   "DB_Integer_IHour" : USInt = PLC Data_Integer.IHour, 1 s
   "DB_Integer_IMinute" : USInt = PLC Data_Integer.IMinute, 1 s
   "DB_Integer_IMonth" : USInt = PLC Data_Integer.IMonth, 1 s
   "DB_Integer_ISecond" : USInt = PLC Data_Integer.ISecond, 1 s
   "DB_Integer_IYear" : UInt = PLC Data_Integer.IYear, 1 s
   "DB_Integer_S1AHour" : USInt = PLC Data_Integer.S1AHour, 1 s
   "DB_Integer_S1AMinute" : USInt = PLC Data_Integer.S1AMinute, 1 s
   "DB_Integer_S1ASecond" : USInt = PLC Data_Integer.S1ASecond, 1 s
   "DB_Integer_S1BHour" : USInt = PLC Data_Integer.S1BHour, 1 s
   "DB_Integer_S1BMinute" : USInt = PLC Data_Integer.S1BMinute, 1 s
   "DB_Integer_S1BSecond" : USInt = PLC Data_Integer.S1BSecond, 1 s
   "DB_Integer_S2AHour" : USInt = PLC Data_Integer.S2AHour, 1 s
   "DB_Integer_S2AMinute" : USInt = PLC Data_Integer.S2AMinute, 1 s
   "DB_Integer_S2ASecond" : USInt = PLC Data_Integer.S2ASecond, 1 s
   "DB_Integer_S2BHour" : USInt = PLC Data_Integer.S2BHour, 1 s
   "DB_Integer_S2BMinute" : USInt = PLC Data_Integer.S2BMinute, 1 s
   "DB_Integer_S2BSecond" : USInt = PLC Data_Integer.S2BSecond, 1 s
   "DB_Integer_S3AHour" : USInt = PLC Data_Integer.S3AHour, 1 s
   "DB_Integer_S3AMinute" : USInt = PLC Data_Integer.S3AMinute, 1 s
   "DB_Integer_S3ASecond" : USInt = PLC Data_Integer.S3ASecond, 1 s
   "DB_Integer_S3BHour" : USInt = PLC Data_Integer.S3BHour, 1 s
   "DB_Integer_S3BMinute" : USInt = PLC Data_Integer.S3BMinute, 1 s
   "DB_Integer_S3BSecond" : USInt = PLC Data_Integer.S3BSecond, 1 s
   "DB_Real_% Reject Out Stop[0]" : Real = PLC Data_Real."% Reject Out Stop"[0], 1 s
   "DB_Real_% Reject Out Stop[1]" : Real = PLC Data_Real."% Reject Out Stop"[1], 1 s
   "DB_Real_% Reject Out Stop[2]" : Real = PLC Data_Real."% Reject Out Stop"[2], 1 s
   "DB_Real_% Reject Out Stop[3]" : Real = PLC Data_Real."% Reject Out Stop"[3], 1 s
   "DB_Real_% Reject Out Stop[4]" : Real = PLC Data_Real."% Reject Out Stop"[4], 1 s
   "DB_Real_% Reject Out Stop[5]" : Real = PLC Data_Real."% Reject Out Stop"[5], 1 s
   "DB_Real_%Bad Read" : Array [0..5] of Real = PLC Data_Real."%Bad Read", 1 s
   "DB_Real_%Bad Read[0]" : Real = PLC Data_Real."%Bad Read"[0], 1 s
   "DB_Real_%Bad Read[1]" : Real = PLC Data_Real."%Bad Read"[1], 1 s
   "DB_Real_%Bad Read[2]" : Real = PLC Data_Real."%Bad Read"[2], 1 s
   "DB_Real_%Bad Read[3]" : Real = PLC Data_Real."%Bad Read"[3], 1 s
   "DB_Real_%Bad Read[4]" : Real = PLC Data_Real."%Bad Read"[4], 1 s
   "DB_Real_%Bad Read[5]" : Real = PLC Data_Real."%Bad Read"[5], 1 s
   "DB_Real_%Good Read[0]" : Real = PLC Data_Real."%Good Read"[0], 1 s
   "DB_Real_%Good Read[1]" : Real = PLC Data_Real."%Good Read"[1], 1 s
   "DB_Real_%Good Read[2]" : Real = PLC Data_Real."%Good Read"[2], 1 s
   "DB_Real_%Good Read[3]" : Real = PLC Data_Real."%Good Read"[3], 1 s
   "DB_Real_%Good Read[4]" : Real = PLC Data_Real."%Good Read"[4], 1 s
   "DB_Real_%Good Read[5]" : Real = PLC Data_Real."%Good Read"[5], 1 s
   "DB_Real_Efficiency CS" : Array [0..5] of Real = PLC Data_Real."% Reject Out Stop", 1 s

discrete alarms
   1: 'Pressure Low', class Errors, trigger "HMI_Tag_1" bit 8
   2: 'Door Open Labelling', class Errors, trigger "HMI_Tag_1" bit 9
   3: 'Door Open Focke Chute', class Errors, trigger "HMI_Tag_1" bit 10
   4: 'Chute 3 Way Full', class Errors, trigger "HMI_Tag_1" bit 11
   5: 'Door Open FC Proximity', class Errors, trigger "HMI_Tag_1" bit 12
   6: 'Alarm2', class Errors, trigger "HMI_Tag_1" bit 13
   7: 'Imaje Paper/Ribbon Out', class Errors, trigger "HMI_Tag_1" bit 14
   8: 'Imaje System Error', class Errors, trigger "HMI_Tag_1" bit 15
   9: 'Imaje Not In Position', class Errors, trigger "HMI_Tag_1" bit 0
   10: 'Heater Not Ready', class Errors, trigger "HMI_Tag_1" bit 1
   11: 'Reed Switch Pneumatic 1 Pusher', class Errors, trigger "HMI_Tag_1" bit 2
   12: 'Alarm3', class Errors, trigger "HMI_Tag_1" bit 3
   13: 'Reed Switch Pneumatic 3 Up', class Errors, trigger "HMI_Tag_1" bit 4
   14: 'Reed Switch Pneumatic 3 Down', class Errors, trigger "HMI_Tag_1" bit 5
   15: 'Reed Switch Pneumatic 4 Down', class Errors, trigger "HMI_Error_Cont" bit 8
   16: 'Reed Switch Pneumatic 4 Up', class Errors, trigger "HMI_Error_Cont" bit 9
   17: 'Reed Switch Pneumatic 5 Advance', class Errors, trigger "HMI_Error_Cont" bit 10
   18: 'Reed Switch Pneumatic 5 Retract', class Errors, trigger "HMI_Error_Cont" bit 11
   19: 'Chute Heating Roll Full', class Errors, trigger "HMI_Tag_1" bit 6

text list "Machine Running": 0 'STOP'; 1 'RUNNING'

text list "Status Markem": 0 'PAUSE'; 1 'START'

text list "Mode Machine": 0 'With Focke Chute'; 1 'Without Focke Chute'

text list "Mode Bypass": 0 'OFF'; 1 'ON'

Template "Template_1" 320x240
   Button "Template_" at 267,190 size 51x47; TextOff 'ExitRuntime'; PictureOff "ExitRuntime_HMI_1"; PictureOn "ExitRuntime_HMI_1"
      on Release: StopRuntime(0)
   Button "Template_1" at 214,190 size 51x47; TextOff 'Text'
   Button "Template_2" at 160,190 size 51x47; TextOff 'Text'
   Button "Template_3" at 107,190 size 51x47; TextOff 'Login'; PictureOff "Login_HMI_1"; PictureOn "Login_HMI_1"
      on Release: function_a2a04561()
   Button "Template_4" at 54,190 size 51x47; TextOff 'AlarmDisplay'; PictureOff "AlarmDisplay_HMI_1"; PictureOn "AlarmDisplay_HMI_1"
      on Release: function_ef3f5d25("Alarm window_Unacknowledged", -1)
   Button "Template_5" at 1,190 size 51x47; TextOff 'NavigateHome'; PictureOff "NavigateHome_HMI_1"; PictureOn "NavigateHome_HMI_1"
   SymbolicIOField "Symbolic_IO_Field_Screen" at 73,7 size 160x25; TextOff '0'; TextOn '1'; TextList "TextList_ScreenNames"
      ProcessValue <- "Tag_ScreenNumber"
   DateTimeField "Template_6" at 235,20 size 85x20
   DateTimeField "Template_7" at 235,0 size 85x20
   GraphicView "Logo" at 0,0 size 71x40; Picture "Logo of HMI_1"

screen "Introduction" 320x240
   Button "Button_1" at 100,200 size 120x30; TextOff 'Go to Main Page'
      on Click: ActivateScreen("Main Page", 0)
   GraphicView "Graphic view_1" at 0,0 size 319x37; Picture "Logo SMS"
   TextField "Text field_1" at 6,54 size 278x31; Text 'END LABELLER MACHINE'
   TextField "Text field_2" at 19,85 size 278x92; Text 'Production : 65 Slof/minute Electric Power : 2,5 KW Compressed Air : 6 Bar Program Version : 14.6 Year : 2013'

screen "Main Page" 320x240
   on GenerateScreen: SetBit("Flag Main Page")
   TextField "Text field_1" at 106,1 size 113x25; Text 'MAIN PAGE'
   TextField "Text field_3" at 5,50 size 91x15; Text 'Machine Status'
   TextField "Text field_4" at 5,73 size 91x15; Text 'Markem Status'
   SymbolicIOField "Symbolic I/O field_2" at 100,48 size 122x19; TextOff '0'; TextOn '1'; TextList "Machine Running"
      ProcessValue <- "Machine Running"
   SymbolicIOField "Symbolic I/O field_1" at 100,71 size 122x19; TextOff '0'; TextOn '1'; TextList "Status Markem"
      ProcessValue <- "Flag Imaje Start"
   Button "Button_4" at 0,209 size 90x30; TextOff 'Test Mode'
      on Click: ActivateScreen("Test Mode", 0)
   Button "Button_5" at 95,209 size 90x30; TextOff 'Parameter'
      on Click: ActivateScreen("Parameter", 0)
   TextField "Text field_5" at 5,95 size 91x15; Text 'Mode Machine'
   SymbolicIOField "Symbolic I/O field_3" at 100,94 size 122x19; TextOff '0'; TextOn '1'; TextList "Mode Machine"
      ProcessValue <- "Flag Enable/Disable Block Focke"
   TextField "Text field_7" at 5,117 size 91x15; Text 'Mode Bypass'
   SymbolicIOField "Symbolic I/O field_4" at 100,117 size 122x19; TextOff '0'; TextOn '1'; TextList "Mode Bypass"
      ProcessValue <- "Flag Machine Bypass"
   IOField "I/O field_3" at 85,24 size 155x23; FormatPattern 9999999999999999999999999999999999999999
      ProcessValue <- "DB_DTL1_Output"
   Button "Button_1" at 287,1 size 29x23; TextOff 'Text'
      on Click: StopRuntime(0)
   Button "Button_2" at 193,208 size 120x30; TextOff 'Statistika Data'
      on Click: ActivateScreen("Data Statistika", 0)

screen "Parameter" 320x240
   on GenerateScreen: SetBit("Flag Parameter Page")
   on ClearScreen: ResetBit("Flag Parameter Page")
   TextField "Text field_1" at 1,0 size 319x27; Text 'PARAMETER'
   Button "Button_4" at 91,202 size 132x30; TextOff 'Back to Main Page'
      on Click: ActivateScreen("Main Page", 0)
   Button "Button_3" at 91,48 size 132x30; TextOff 'Setting Timer'
      on Click: ActivateScreen("Setting Timer", 0)
   Button "Button_2" at 91,88 size 132x30; TextOff 'Setting Machine'
      on Click: ActivateScreen("Setting Machine", 0)

screen "Setting Timer" 320x240
   on ClearScreen: ResetBit("Flag Parameter Page")
   on GenerateScreen: SetBit("Flag Parameter Page")
   TextField "Text field_1" at 0,0 size 319x27; Text 'SETTING TIMER'
   Button "Button_2" at 92,200 size 120x30; TextOff 'Back to Parameter'
      on Click: ActivateScreen("Parameter", 0)
   TextField "Text field_2" at 5,39 size 150x15; Text 'Timer Delay Stamp'
   IOField "I/O field_1" at 152,40 size 80x16; FormatPattern 9999; Unit  ms
      ProcessValue <- "Timer Delay Stamp"
   TextField "Text field_3" at 5,63 size 150x15; Text 'Timer Scanning Barcode'
   IOField "I/O field_2" at 153,64 size 80x16; FormatPattern 9999; Unit  ms
      ProcessValue <- "Timer Trigger Barcode"

screen "Test Mode" 320x240
   on GenerateScreen: SetBit("PB Test Mode")
   on ClearScreen: ResetBit("PB Test Mode")
   TextField "Text field_1" at 1,1 size 319x27; Text 'TEST MODE'
   Switch "Switch_1" at 3,34 size 95x30; TextOff 'Pneumatic 1 Off'; CaptionText 'Switch'; TextOn 'Pneumatic 1 On'
      ProcessValue <- "PB Test Pneumatic 1"
   Switch "Switch_2" at 3,75 size 95x30; CaptionText 'Switch'; TextOff 'Pneumatic 2 Off'; TextOn 'Pneumatic 2 On'
      ProcessValue <- "PB Test Pneumatic 2"
   Switch "Switch_3" at 3,116 size 95x30; CaptionText 'Switch'; TextOff 'Pneumatic 3 Off'; TextOn 'Pneumatic 3 On'
      ProcessValue <- "PB Test Pneumatic 3"
   Switch "Switch_5" at 104,34 size 115x30; CaptionText 'Switch'; TextOff 'Pneumatic 5 Off'; TextOn 'Pneumatic 5 On'
      ProcessValue <- "PB Test Pneumatic 5"
   Switch "Switch_6" at 226,116 size 90x30; CaptionText 'Switch'; TextOff 'Motor Off'; TextOn 'Motor On'
      ProcessValue <- "PB Test Motor"
   Button "Button_1" at 100,204 size 120x30; TextOff 'Back to Main Page'
      on Click: ActivateScreen("Main Page", 0)
   Button "Button_2" at 226,34 size 90x30; TextOff 'Stamp Off'; TextOn 'Stamp On'
      on Press: SetBit("PB Test Imaje")
      on Release: ResetBit("PB Test Imaje")
   Switch "Switch_7" at 104,116 size 115x30; CaptionText 'Switch'; TextOff 'Air Valve On'; TextOn 'Air Valve Off'
      ProcessValue <- "PB Test Air Valve"
   Button "Button_3" at 226,75 size 90x30; TextOff 'Teach In'
      on Press: SetBit("Flag Teach In Barcode")
      on Release: ResetBit("Flag Teach In Barcode")
   Switch "Switch_8" at 3,157 size 95x30; CaptionText 'Switch'; TextOff 'Pneumatic 4 Off'; TextOn 'Pneumatic 4 On'
      ProcessValue <- "PB Test Pneumatic 4"
   Switch "Switch_4" at 104,75 size 115x30; CaptionText 'Switch'; TextOff 'Pneumatic 6 On'; TextOn 'Pneumatic 6 Off'
      ProcessValue <- "PB Test Pneumatic 6"
   Switch "Switch_9" at 104,157 size 115x30; CaptionText 'Switch'; TextOff 'Conveyor Pusher Off'; TextOn 'Conveyor Pusher On'
      ProcessValue <- "PB Test Motor Coveyor Pusher"
   Switch "Switch_10" at 226,157 size 90x30; CaptionText 'Switch'; TextOff 'Heating Roll Off'; TextOn 'Heating Roll On'
      ProcessValue <- "PB Test Motor Heating Roll"

screen "Setting Machine" 320x240
   on ClearScreen: ResetBit("Flag Parameter Page")
   on GenerateScreen: SetBit("Flag Parameter Page")
   TextField "Text field_1" at 1,0 size 319x27; Text 'SETTING MACHINE'
   Switch "Switch_1" at 16,38 size 135x30; CaptionText 'Switch'; TextOff 'Barcode Off'; TextOn 'Barcode ON'
      ProcessValue <- "Flag Barcode HMI"
   Switch "Switch_2" at 16,108 size 135x30; CaptionText 'Switch'; TextOff 'Chute 3Way Error ON'; TextOn 'Chute 3Way Error OFF'
      ProcessValue <- "Flag Enable/Disable Error Chute 3 Way"
   Button "Button_2" at 101,205 size 120x30; TextOff 'Back to Parameter'
      on Click: ActivateScreen("Parameter", 0)
   Switch "Switch_3" at 16,73 size 135x30; CaptionText 'Switch'; TextOff 'Heater Error Off'; TextOn 'Heater Error ON'
      ProcessValue <- "Flag Heater Error HMI"
   Switch "Switch_4" at 170,38 size 135x30; CaptionText 'Switch'; TextOff 'Reed Switch Bypass Off'; TextOn 'Reed Switch Bypass On'
      ProcessValue <- "Flag Pneumatic Bypass"
   Switch "Switch_5" at 170,108 size 135x30; CaptionText 'Switch'; TextOff 'Safety Door On'; TextOn 'Safety Door Off'
      ProcessValue <- "Flag Enable/Disable Error Door Open"
   Button "Button_1" at 289,0 size 31x30; TextOff 'Setting Mode'; Authorization "User administration"
      on Click: ActivateScreen("Setting Mode", 0)
   Button "Button_3" at 170,73 size 135x30; TextOff 'Setting Reed Switch'
      on Click: ActivateScreen("Setting Reed Switch", 0)
   Switch "Switch_6" at 16,143 size 135x30; CaptionText 'Switch'; TextOff 'Chute Heating Roll Error ON'; TextOn 'Chute Heating Roll Error OFF'
      ProcessValue <- "Flag Enable/Disable Error Chute Before Heating Roll"
   Softkey "Softkey_F6" at 266,202 size 53x38
      on KeyDown: ActivateScreen("Setting Mode", 0)
      on KeyUp: ActivateScreen("Setting Mode", 0)
   Softkey "Softkey_F5" at 213,202 size 53x38
      on KeyDown: function_f23ef4c9()
      on KeyUp: function_f23ef4c9()

screen "Setting Mode" 320x240
   TextField "Text field_1" at 1,0 size 319x27; Text 'MODE MACHINE'
   Button "Button_1" at 95,203 size 129x30; TextOff 'Back to Setting Machine'
      on Click: ActivateScreen("Setting Machine", 0)
   Switch "Switch_1" at 70,46 size 177x32; CaptionText 'Switch'; TextOff 'With Focke Chute'; TextOn 'Without Focke Chute'
      ProcessValue <- "Flag Enable/Disable Block Focke"
   Switch "Switch_2" at 70,90 size 177x32; TextOff 'Disable Flow to Reject'; CaptionText 'Switch'; TextOn 'Enable Flow to Reject'
      ProcessValue <- "Flag Enable/Disable Flow to Reject"
   Switch "Switch_3" at 70,130 size 177x32; TextOff 'With Heating Roll'; CaptionText 'Switch'; TextOn 'Without Heating Roll'
      ProcessValue <- "Flag Enable/Disable Heating Roll"

screen "Setting Reed Switch" 320x240
   TextField "Text field_1" at 1,3 size 319x27; Text 'SETTING REED SWITCH BYPASS'
   Switch "Switch_4" at 21,103 size 128x30; CaptionText 'Switch'; TextOff 'RS Pneu 3 Bypass Off'; TextOn 'RS Pneu 3 Bypass On'
      ProcessValue <- "RS Bypass Pneumatic 3"
   Switch "Switch_1" at 172,103 size 128x30; CaptionText 'Switch'; TextOff 'RS Pneu 5 Bypass Off'; TextOn 'RS Pneu 5 Bypass On'
      ProcessValue <- "RS Bypass Pneumatic 5"
   Switch "Switch_2" at 172,59 size 128x30; CaptionText 'Switch'; TextOff 'RS Pneu 4 Bypass Off'; TextOn 'RS Pneu 4 Bypass On'
      ProcessValue <- "RS Bypass Pneumatic 4"
   Switch "Switch_3" at 21,59 size 128x30; CaptionText 'Switch'; TextOff 'RS Pneu 1 Bypass Off'; TextOn 'RS Pneu 1 Bypass On'
      ProcessValue <- "RS Bypass Pneumatic 1"
   Button "Button_1" at 95,203 size 129x30; TextOff 'Back to Setting Machine'
      on Click: ActivateScreen("Setting Machine", 0)

screen "Data Current Shift" 320x240
   IOField "I/O field_11" at 221,82 size 60x19; FormatPattern 999.99; Unit   %
      ProcessValue <- "Data_Real_% Total Output[0]"
   IOField "I/O field_9" at 221,102 size 60x19; FormatPattern 999.99; Unit   %
      ProcessValue <- "DB_Real_%Good Read[0]"
   IOField "I/O field_8" at 221,120 size 60x19; FormatPattern 999.99; Unit   %
      ProcessValue <- "DB_Real_%Bad Read[0]"
   TextField "Text field_1" at 92,0 size 137x18; Text 'CURRENT SHIFT DATA'
   IOField "I/O field_1" at 142,59 size 79x19; FormatPattern 99999999; Unit  Pcs
      ProcessValue <- "DB_IntData_Input Sloft"
   TextField "Text field_2" at 4,60 size 138x17; Text 'Input Sloft'
   TextField "Text field_3" at 4,83 size 138x17; Text 'Total Output Sloft'
   TextField "Text field_4" at 4,101 size 138x19; Text 'Good Read Sloft'
   TextField "Text field_7" at 4,121 size 138x18; Text 'Bad Read Sloft'
   IOField "I/O field_3" at 142,101 size 79x19; FormatPattern 99999999; Unit  Pcs
      ProcessValue <- "DB_IntData_Good R1"
   IOField "I/O field_5" at 142,82 size 79x22; FormatPattern 99999999; Unit  Pcs
      ProcessValue <- "DB_IntData_Tot Good R"
   IOField "I/O field_4" at 142,121 size 79x18; FormatPattern 99999999; Unit  Pcs
      ProcessValue <- "DB_IntData_Bad R"
   IOField "I/O field_6" at 4,32 size 132x18; FormatPattern 9999999999999999999999999999999999999999
      ProcessValue <- "DB_DTL1_Cur_ShiftA"
   TextField "Text field_9" at 142,31 size 19x15; Text 'S/D'
   Button "Button_1" at 52,206 size 90x32; TextOff 'Back To Statistika Data'; TextOn 'Statistika Data'
      on Click: ActivateScreen("Data Statistika", 0)
   Button "Button_3" at 4,205 size 41x34; TextOff 'Main Page'; PictureOff "Home"
      on Click: ActivateScreen("Main Page", 0)
   Button "Button_2" at 226,207 size 90x30; TextOff 'Next Data --->'; TextOn 'Error Counter'
      on Click: ActivateScreen("Data Time Current Shift", 0)
   IOField "I/O field_7" at 167,32 size 132x18; FormatPattern 9999999999999999999999999999999999999999
      ProcessValue <- "DB_DTL1_Cur_ShiftB"

screen "Data Current Shift_1" 320x240
   IOField "I/O field_11" at 221,82 size 60x19; FormatPattern 999.99; Unit   %
      ProcessValue <- "Data_Real_% Total Output[1]"
   IOField "I/O field_8" at 221,118 size 60x19; FormatPattern 999.99; Unit   %
      ProcessValue <- "DB_Real_%Bad Read[1]"
   IOField "I/O field_9" at 221,101 size 60x19; FormatPattern 999.99; Unit   %
      ProcessValue <- "DB_Real_%Good Read[1]"
   TextField "Text field_1" at 67,1 size 193x18; Text 'CURRENT SHIFT DATA MINUS 1'
   IOField "I/O field_1" at 142,59 size 79x19; FormatPattern 99999999; Unit  Pcs
      ProcessValue <- "DB_IntData_Input Sloft_1"
   TextField "Text field_2" at 4,60 size 138x17; Text 'Input Sloft'
   Button "Button_1" at 55,203 size 90x32; TextOff 'Back To Statistika Data'; TextOn 'Statistika Data'
      on Click: ActivateScreen("Data Statistika", 0)
   Button "Button_3" at 4,202 size 45x34; TextOff 'Main Page'; PictureOff "Home"
      on Click: ActivateScreen("Main Page", 0)
   Button "Button_2" at 223,205 size 90x30; TextOff 'Next Data --->'; TextOn 'Error Counter'
      on Click: ActivateScreen("Data Time Current Shift_1", 0)
   IOField "I/O field_6" at 4,32 size 132x18; FormatPattern 9999999999999999999999999999999999999999
      ProcessValue <- "DB_DTL1_Cur_ShiftA_1"
   TextField "Text field_9" at 142,31 size 19x15; Text 'S/D'
   IOField "I/O field_7" at 167,32 size 132x18; FormatPattern 9999999999999999999999999999999999999999
      ProcessValue <- "DB_DTL1_Cur_ShiftB_1"
   TextField "Text field_3" at 4,83 size 138x17; Text 'Total Output Sloft'
   TextField "Text field_4" at 4,101 size 138x19; Text 'Good Read Sloft'
   TextField "Text field_7" at 4,119 size 138x18; Text 'Bad Read Sloft'
   IOField "I/O field_3" at 142,101 size 79x19; FormatPattern 9999999999; Unit  Pcs
      ProcessValue <- "DB_IntData_Good R1_1"
   IOField "I/O field_5" at 142,82 size 79x22; FormatPattern 99999999; Unit  Pcs
      ProcessValue <- "DB_IntData_Tot Out Slof_1"
   IOField "I/O field_4" at 142,119 size 79x18; FormatPattern 9999999999; Unit  Pcs
      ProcessValue <- "DB_IntData_Bad R_1"

screen "Data Current Shift_2" 320x240
   IOField "I/O field_11" at 221,82 size 60x19; FormatPattern 999.99; Unit   %
      ProcessValue <- "Data_Real_% Total Output[2]"
   IOField "I/O field_8" at 222,119 size 60x19; FormatPattern 999.99; Unit   %
      ProcessValue <- "DB_Real_%Bad Read[2]"
   IOField "I/O field_9" at 221,100 size 60x19; FormatPattern 999.99; Unit   %
      ProcessValue <- "DB_Real_%Good Read[2]"
   TextField "Text field_1" at 67,1 size 193x18; Text 'CURRENT SHIFT DATA MINUS 2'
   IOField "I/O field_1" at 142,59 size 79x19; FormatPattern 99999999; Unit  Pcs
      ProcessValue <- "DB_IntData_Input Sloft_2"
   TextField "Text field_2" at 4,60 size 138x17; Text 'Input Sloft'
   Button "Button_1" at 57,204 size 90x32; TextOff 'Back To Statistika Data'; TextOn 'Statistika Data'
      on Click: ActivateScreen("Data Statistika", 0)
   Button "Button_3" at 4,202 size 45x34; TextOff 'Main Page'; PictureOff "Home"
      on Click: ActivateScreen("Main Page", 0)
   Button "Button_2" at 221,206 size 90x30; TextOff 'Next Data --->'; TextOn 'Error Counter'
      on Click: ActivateScreen("Data Time Current Shift_2", 0)
   IOField "I/O field_6" at 4,32 size 132x18; FormatPattern 9999999999999999999999999999999999999999
      ProcessValue <- "DB_DTL1_Cur_ShiftA_2"
   TextField "Text field_9" at 142,31 size 19x15; Text 'S/D'
   IOField "I/O field_7" at 167,32 size 132x18; FormatPattern 9999999999999999999999999999999999999999
      ProcessValue <- "DB_DTL1_Cur_ShiftB_2"
   TextField "Text field_3" at 4,83 size 138x17; Text 'Total Output Sloft'
   TextField "Text field_4" at 4,101 size 138x19; Text 'Good Read Sloft'
   TextField "Text field_7" at 5,120 size 138x18; Text 'Bad Read Sloft'
   IOField "I/O field_3" at 142,101 size 79x19; FormatPattern 9999999999; Unit  Pcs
      ProcessValue <- "DB_IntData_Good R1_2"
   IOField "I/O field_5" at 142,82 size 79x22; FormatPattern 9999999999; Unit  Pcs
      ProcessValue <- "DB_IntData_Tot Good R_2"
   IOField "I/O field_4" at 143,120 size 79x18; FormatPattern 9999999999; Unit  Pcs
      ProcessValue <- "DB_IntData_Bad R_2"

screen "Data Current Shift_3" 320x240
   IOField "I/O field_11" at 221,83 size 60x19; FormatPattern 999.99; Unit   %
      ProcessValue <- "Data_Real_% Total Output[3]"
   IOField "I/O field_8" at 221,119 size 60x19; FormatPattern 999.99; Unit   %
      ProcessValue <- "DB_Real_%Bad Read[3]"
   IOField "I/O field_9" at 221,100 size 60x19; FormatPattern 999.99; Unit   %
      ProcessValue <- "DB_Real_%Good Read[3]"
   TextField "Text field_1" at 67,1 size 193x18; Text 'CURRENT SHIFT DATA MINUS 3'
   IOField "I/O field_1" at 142,59 size 79x19; FormatPattern 99999999; Unit  Pcs
      ProcessValue <- "DB_IntData_Input Sloft_3"
   TextField "Text field_2" at 4,60 size 138x17; Text 'Input Sloft'
   Button "Button_1" at 58,205 size 90x32; TextOff 'Back To Statistika Data'; TextOn 'Statistika Data'
      on Click: ActivateScreen("Data Statistika", 0)
   Button "Button_3" at 6,203 size 45x34; TextOff 'Main Page'; PictureOff "Home"
      on Click: ActivateScreen("Main Page", 0)
   Button "Button_2" at 221,206 size 90x30; TextOff 'Next Data --->'; TextOn 'Error Counter'
      on Click: ActivateScreen("Data Time Current Shift_3", 0)
   IOField "I/O field_6" at 4,32 size 132x18; FormatPattern 9999999999999999999999999999999999999999
      ProcessValue <- "DB_DTL1_Cur_ShiftA_3"
   TextField "Text field_9" at 142,31 size 19x15; Text 'S/D'
   IOField "I/O field_7" at 167,32 size 132x18; FormatPattern 9999999999999999999999999999999999999999
      ProcessValue <- "DB_DTL1_Cur_ShiftB_3"
   TextField "Text field_3" at 4,83 size 138x17; Text 'Total Output Sloft'
   TextField "Text field_4" at 4,101 size 138x19; Text 'Good Read Sloft'
   TextField "Text field_7" at 4,120 size 138x18; Text 'Bad Read Sloft'
   IOField "I/O field_3" at 142,101 size 79x19; FormatPattern 9999999999; Unit  Pcs
      ProcessValue <- "DB_IntData_Good R1_3"
   IOField "I/O field_5" at 142,82 size 79x22; FormatPattern 9999999999; Unit  Pcs
      ProcessValue <- "DB_IntData_Tot Good R_3"
   IOField "I/O field_4" at 142,120 size 79x18; FormatPattern 9999999999; Unit  Pcs
      ProcessValue <- "DB_IntData_Bad R_3"

screen "Data Current Shift_4" 320x240
   IOField "I/O field_11" at 223,82 size 60x19; FormatPattern 999.99; Unit   %
      ProcessValue <- "Data_Real_% Total Output[4]"
   IOField "I/O field_8" at 222,119 size 60x19; FormatPattern 999.99; Unit   %
      ProcessValue <- "DB_Real_%Bad Read[4]"
   IOField "I/O field_9" at 222,100 size 60x19; FormatPattern 999.99; Unit   %
      ProcessValue <- "DB_Real_%Good Read[4]"
   TextField "Text field_1" at 67,1 size 193x18; Text 'CURRENT SHIFT DATA MINUS 4'
   IOField "I/O field_1" at 142,59 size 79x19; FormatPattern 99999999; Unit  Pcs
      ProcessValue <- "DB_IntData_Input Sloft_4"
   TextField "Text field_2" at 4,60 size 138x17; Text 'Input Sloft'
   Button "Button_1" at 56,205 size 90x32; TextOff 'Back To Statistika Data'; TextOn 'Statistika Data'
      on Click: ActivateScreen("Data Statistika", 0)
   Button "Button_3" at 4,203 size 45x34; TextOff 'Main Page'; PictureOff "Home"
      on Click: ActivateScreen("Main Page", 0)
   Button "Button_2" at 216,206 size 90x30; TextOff 'Next Data --->'; TextOn 'Error Counter'
      on Click: ActivateScreen("Data Time Current Shift_4", 0)
   IOField "I/O field_6" at 4,32 size 132x18; FormatPattern 9999999999999999999999999999999999999999
      ProcessValue <- "DB_DTL1_Cur_ShiftA_4"
   TextField "Text field_9" at 142,31 size 19x15; Text 'S/D'
   IOField "I/O field_7" at 167,32 size 132x18; FormatPattern 9999999999999999999999999999999999999999
      ProcessValue <- "DB_DTL1_Cur_ShiftB_4"
   TextField "Text field_3" at 4,83 size 138x17; Text 'Total Output Sloft'
   TextField "Text field_4" at 4,101 size 138x19; Text 'Good Read Sloft'
   TextField "Text field_7" at 4,120 size 138x18; Text 'Bad Read Sloft'
   IOField "I/O field_3" at 142,101 size 79x19; FormatPattern 9999999999; Unit  Pcs
      ProcessValue <- "DB_IntData_Good R1_4"
   IOField "I/O field_5" at 142,82 size 79x22; FormatPattern 9999999999; Unit  Pcs
      ProcessValue <- "DB_IntData_Tot Good R_4"
   IOField "I/O field_4" at 142,120 size 79x18; FormatPattern 9999999999; Unit  Pcs
      ProcessValue <- "DB_IntData_Bad R_4"

screen "Data Current Shift_5" 320x240
   IOField "I/O field_11" at 221,82 size 60x19; FormatPattern 999.99; Unit   %
      ProcessValue <- "Data_Real_% Total Output[5]"
   IOField "I/O field_8" at 221,119 size 60x19; FormatPattern 999.99; Unit   %
      ProcessValue <- "DB_Real_%Bad Read[5]"
   IOField "I/O field_9" at 221,100 size 60x19; FormatPattern 999.99; Unit   %
      ProcessValue <- "DB_Real_%Good Read[5]"
   TextField "Text field_1" at 67,1 size 193x18; Text 'CURRENT SHIFT DATA MINUS 5'
   IOField "I/O field_1" at 142,59 size 79x19; FormatPattern 99999999; Unit  Pcs
      ProcessValue <- "DB_IntData_Input Sloft_5"
   TextField "Text field_2" at 4,60 size 138x17; Text 'Input Sloft'
   Button "Button_1" at 59,203 size 90x32; TextOff 'Back To Statistika Data'; TextOn 'Statistika Data'
      on Click: ActivateScreen("Data Statistika", 0)
   Button "Button_3" at 7,202 size 45x34; TextOff 'Main Page'; PictureOff "Home"
      on Click: ActivateScreen("Main Page", 0)
   Button "Button_2" at 219,204 size 90x30; TextOff 'Next Data --->'; TextOn 'Error Counter'
      on Click: ActivateScreen("Data Current Shift_5", 0)
   IOField "I/O field_6" at 4,32 size 132x18; FormatPattern 9999999999999999999999999999999999999999
      ProcessValue <- "DB_DTL1_Cur_ShiftA_5"
   TextField "Text field_9" at 142,31 size 19x15; Text 'S/D'
   IOField "I/O field_7" at 167,32 size 132x18; FormatPattern 9999999999999999999999999999999999999999
      ProcessValue <- "DB_DTL1_Cur_ShiftB_5"
   TextField "Text field_3" at 4,83 size 138x17; Text 'Total Output Sloft'
   TextField "Text field_4" at 4,101 size 138x19; Text 'Good Read Sloft'
   TextField "Text field_7" at 4,120 size 138x18; Text 'Bad Read Sloft'
   IOField "I/O field_3" at 142,101 size 79x19; FormatPattern 9999999999; Unit  Pcs
      ProcessValue <- "DB_IntData_Good R1_5"
   IOField "I/O field_5" at 142,82 size 79x22; FormatPattern 9999999999; Unit  Pcs
      ProcessValue <- "DB_IntData_Tot Good R_5"
   IOField "I/O field_4" at 142,120 size 79x18; FormatPattern 9999999999; Unit  Pcs
      ProcessValue <- "DB_IntData_Bad R_5"

screen "Data Statistika" 320x240
   Button "Button_1" at 9,47 size 146x30; TextOff 'Current Shift Data'
      on Click: ActivateScreen("Data Current Shift", 0)
   Button "Button_2" at 284,3 size 27x24; TextOff 'Text'; TextOn 'Statistik Parameter'; Authorization "User administration"
      on Click: ActivateScreen("Statistik Parameter", 0)
   Button "Button_3" at 9,80 size 146x30; TextOff 'Current Shift Data Minus 1'
      on Click: ActivateScreen("Data Current Shift_1", 0)
   Button "Button_4" at 9,113 size 147x30; TextOff 'Current Shift Data Minus 2'
      on Click: ActivateScreen("Data Current Shift_2", 0)
   Button "Button_5" at 163,46 size 147x30; TextOff 'Current Shift Data Minus 3'
      on Click: ActivateScreen("Data Current Shift_3", 0)
   Button "Button_6" at 163,80 size 147x30; TextOff 'Current Shift Data Minus 4'
      on Click: ActivateScreen("Data Current Shift_4", 0)
   Button "Button_7" at 163,113 size 147x30; TextOff 'Current Shift Data Minus 5'
      on Click: ActivateScreen("Data Current Shift_5", 0)
   TextField "Text field_1" at 99,4 size 106x18; Text 'STATISTIC DATA'
   Button "Button_8" at 91,209 size 132x30; TextOff 'Back to Main Page'
      on Click: ActivateScreen("Main Page", 0)

screen "Error Counter" 320x240
   TextField "Text field_34" at 6,153 size 21x19; Text '6'
   TextField "Text field_33" at 7,133 size 21x19; Text '5'
   TextField "Text field_32" at 7,114 size 21x19; Text '4'
   TextField "Text field_31" at 7,95 size 21x19; Text '3'
   TextField "Text field_30" at 7,76 size 21x19; Text '2'
   TextField "Text field_29" at 7,58 size 21x19; Text '1'
   TextField "Text field_28" at 7,40 size 21x19; Text 'No'
   IOField "I/O field_8" at 225,153 size 26x19; FormatPattern 999
      ProcessValue <- "DB_DTLData_DTL_RS Pneu Er.SECOND"
   IOField "I/O field_16" at 200,153 size 25x19; FormatPattern 999
      ProcessValue <- "DB_DTLData_DTL_RS Pneu Er.MINUTE"
   IOField "I/O field_17" at 175,153 size 25x19; FormatPattern 999
      ProcessValue <- "DB_DTLData_DTL_RS Pneu Er.HOUR"
   TextField "Text field_8" at 29,153 size 145x19; Text 'Reed Swicth Pneumatic Error'
   TextField "Text field_10" at 196,152 size 8x17; Text ':'
   TextField "Text field_21" at 220,153 size 8x17; Text ':'
   IOField "I/O field_21" at 225,94 size 26x19; FormatPattern 999
      ProcessValue <- "Data_DTLData_DTL_Imaje Not In Position[0].SECOND"
   IOField "I/O field_22" at 200,94 size 25x19; FormatPattern 999
      ProcessValue <- "Data_DTLData_DTL_Imaje Not In Position[0].MINUTE"
   IOField "I/O field_23" at 175,94 size 25x19; FormatPattern 999
      ProcessValue <- "Data_DTLData_DTL_Imaje Not In Position[0].HOUR"
   TextField "Text field_25" at 29,95 size 145x19; Text 'Imaje Not In Position'
   IOField "I/O field_18" at 225,76 size 26x19; FormatPattern 999
      ProcessValue <- "Data_DTLData_DTL_Paper R Out[0].SECOND"
   IOField "I/O field_19" at 200,76 size 25x19; FormatPattern 999
      ProcessValue <- "Data_DTLData_DTL_Paper R Out[0].MINUTE"
   IOField "I/O field_20" at 175,76 size 25x19; FormatPattern 999
      ProcessValue <- "Data_DTLData_DTL_Paper R Out[0].HOUR"
   TextField "Text field_22" at 29,76 size 145x19; Text 'Imaje Papper Or Ribbon Out'
   TextField "Text field_2" at 176,43 size 24x15; Text 'Hour'
   IOField "I/O field_10" at 225,134 size 26x19; FormatPattern 999
      ProcessValue <- "DB_DTLData_DTL_Slof Jam.SECOND"
   IOField "I/O field_11" at 200,134 size 25x19; FormatPattern 999
      ProcessValue <- "DB_DTLData_DTL_Slof Jam.MINUTE"
   IOField "I/O field_12" at 175,134 size 25x19; FormatPattern 999
      ProcessValue <- "DB_DTLData_DTL_Slof Jam.HOUR"
   IOField "I/O field_4" at 225,114 size 26x19; FormatPattern 999
      ProcessValue <- "DB_DTLData_DTL_Press Low.SECOND"
   IOField "I/O field_5" at 200,114 size 25x19; FormatPattern 999
      ProcessValue <- "DB_DTLData_DTL_Press Low.MINUTE"
   IOField "I/O field_9" at 175,114 size 25x19; FormatPattern 999
      ProcessValue <- "DB_DTLData_DTL_Press Low.HOUR"
   TextField "Text field_12" at 229,43 size 19x15; Text 'Sec'
   TextField "Text field_11" at 203,43 size 19x15; Text 'Min'
   IOField "I/O field_2" at 225,59 size 26x19; FormatPattern 999
      ProcessValue <- "DB_DTLData_DTL_Imaje Er.SECOND"
   IOField "I/O field_1" at 200,59 size 25x19; FormatPattern 999
      ProcessValue <- "DB_DTLData_DTL_Imaje Er.MINUTE"
   TextField "Text field_1" at 54,1 size 213x18; Text 'CURRENT SHIFT DATA (Detil Error)'
   TextField "Text field_3" at 30,42 size 144x17; Text 'Error Counter'
   TextField "Text field_4" at 29,59 size 145x19; Text 'System Imaje Error'
   TextField "Text field_5" at 29,114 size 145x21; Text 'Pressure Low'
   TextField "Text field_6" at 29,133 size 145x20; Text 'Sloft Jammed'
   IOField "I/O field_3" at 175,59 size 25x19; FormatPattern 999
      ProcessValue <- "DB_DTLData_DTL_Imaje Er.HOUR"
   TextField "Text field_13" at 196,58 size 8x17; Text ':'
   TextField "Text field_14" at 196,113 size 8x17; Text ':'
   TextField "Text field_15" at 196,133 size 8x17; Text ':'
   TextField "Text field_17" at 220,58 size 8x17; Text ':'
   TextField "Text field_18" at 220,113 size 8x17; Text ':'
   TextField "Text field_19" at 220,133 size 8x17; Text ':'
   Button "Button_3" at 5,203 size 45x34; TextOff 'Main Page'; PictureOff "Home"
      on Click: ActivateScreen("Main Page", 0)
   Button "Button_1" at 54,209 size 93x28; TextOff 'Back To Data Statistika'; TextOn 'Data Statistika'
      on Click: ActivateScreen("Data Statistika", 0)
   Button "Button_2" at 219,209 size 97x28; TextOff '<----- Back'; TextOn 'Sloft Data'
      on Click: ActivateScreen("Data Time Current Shift", 0)
   IOField "I/O field_6" at 6,19 size 132x18; FormatPattern 9999999999999999999999999999999999999999
      ProcessValue <- "DB_DTL1_Cur_ShiftA"
   TextField "Text field_9" at 145,19 size 19x15; Text 'S/D'
   IOField "I/O field_7" at 169,18 size 127x17; FormatPattern 9999999999999999999999999999999999999999
      ProcessValue <- "DB_DTL1_Cur_ShiftB"
   TextField "Text field_23" at 196,75 size 8x17; Text ':'
   TextField "Text field_24" at 220,75 size 8x17; Text ':'
   TextField "Text field_26" at 196,93 size 8x17; Text ':'
   TextField "Text field_27" at 220,93 size 8x17; Text ':'

screen "Error Counter_1" 320x240
   TextField "Text field_1" at 24,1 size 269x18; Text 'CURRENT SHIFT DATA MINUS 1 (Detil Error)'
   Button "Button_3" at 0,200 size 45x34; TextOff 'Main Page'; PictureOff "Home"
      on Click: ActivateScreen("Main Page", 0)
   Button "Button_1" at 52,206 size 93x28; TextOff 'Back To Data Statistika'; TextOn 'Data Statistika'
      on Click: ActivateScreen("Data Statistika", 0)
   Button "Button_2" at 207,206 size 97x28; TextOff '<----- Back'; TextOn 'Sloft Data'
      on Click: ActivateScreen("Data Time Current Shift_1", 0)
   IOField "I/O field_6" at 6,19 size 132x18; FormatPattern 9999999999999999999999999999999999999999
      ProcessValue <- "DB_DTL1_Cur_ShiftA_1"
   TextField "Text field_9" at 145,20 size 19x15; Text 'S/D'
   IOField "I/O field_7" at 169,20 size 132x18; FormatPattern 9999999999999999999999999999999999999999
      ProcessValue <- "DB_DTL1_Cur_ShiftB_1"
   TextField "Text field_34" at 6,153 size 21x19; Text '6'
   TextField "Text field_33" at 7,133 size 21x19; Text '5'
   TextField "Text field_32" at 7,114 size 21x19; Text '4'
   TextField "Text field_31" at 7,95 size 21x19; Text '3'
   TextField "Text field_30" at 7,76 size 21x19; Text '2'
   TextField "Text field_29" at 7,58 size 21x19; Text '1'
   TextField "Text field_28" at 7,40 size 21x19; Text 'No'
   IOField "I/O field_8" at 225,153 size 26x19; FormatPattern 999
      ProcessValue <- "DB_DTLData_DTL_RS Pneu Er_1.SECOND"
   IOField "I/O field_16" at 200,153 size 25x19; FormatPattern 999
      ProcessValue <- "DB_DTLData_DTL_RS Pneu Er_1.MINUTE"
   IOField "I/O field_17" at 175,153 size 25x19; FormatPattern 999
      ProcessValue <- "DB_DTLData_DTL_RS Pneu Er_1.HOUR"
   TextField "Text field_8" at 29,153 size 145x19; Text 'Reed Swicth Pneumatic Error'
   TextField "Text field_10" at 196,152 size 8x17; Text ':'
   TextField "Text field_21" at 220,153 size 8x17; Text ':'
   IOField "I/O field_21" at 225,94 size 26x19; FormatPattern 999
      ProcessValue <- "Data_DTLData_DTL_Imaje Not In Position[1].SECOND"
   IOField "I/O field_22" at 200,94 size 25x19; FormatPattern 999
      ProcessValue <- "Data_DTLData_DTL_Imaje Not In Position[1].MINUTE"
   IOField "I/O field_23" at 175,94 size 25x19; FormatPattern 999
      ProcessValue <- "Data_DTLData_DTL_Imaje Not In Position[1].HOUR"
   TextField "Text field_25" at 29,95 size 145x19; Text 'Imaje Not In Position'
   IOField "I/O field_18" at 225,76 size 26x19; FormatPattern 999
      ProcessValue <- "Data_DTLData_DTL_Paper R Out[1].SECOND"
   IOField "I/O field_19" at 200,76 size 25x19; FormatPattern 999
      ProcessValue <- "Data_DTLData_DTL_Paper R Out[1].MINUTE"
   IOField "I/O field_20" at 175,76 size 25x19; FormatPattern 999
      ProcessValue <- "Data_DTLData_DTL_Paper R Out[1].HOUR"
   TextField "Text field_22" at 29,76 size 145x19; Text 'Imaje Papper Or Ribbon Out'
   TextField "Text field_2" at 176,43 size 24x15; Text 'Hour'
   IOField "I/O field_10" at 225,134 size 26x19; FormatPattern 999
      ProcessValue <- "DB_DTLData_DTL_Slof Jam_1.SECOND"
   IOField "I/O field_11" at 200,134 size 25x19; FormatPattern 999
      ProcessValue <- "DB_DTLData_DTL_Slof Jam_1.MINUTE"
   IOField "I/O field_12" at 175,134 size 25x19; FormatPattern 999
      ProcessValue <- "DB_DTLData_DTL_Slof Jam_1.HOUR"
   IOField "I/O field_4" at 225,114 size 26x19; FormatPattern 999
      ProcessValue <- "DB_DTLData_DTL_Press Low_1.SECOND"
   IOField "I/O field_5" at 200,114 size 25x19; FormatPattern 999
      ProcessValue <- "DB_DTLData_DTL_Press Low_1.MINUTE"
   IOField "I/O field_9" at 175,114 size 25x19; FormatPattern 999
      ProcessValue <- "DB_DTLData_DTL_Press Low_1.HOUR"
   TextField "Text field_12" at 229,43 size 19x15; Text 'Sec'
   TextField "Text field_11" at 203,43 size 19x15; Text 'Min'
   IOField "I/O field_2" at 225,59 size 26x19; FormatPattern 999
      ProcessValue <- "DB_DTLData_DTL_Imaje Er_1.SECOND"
   IOField "I/O field_1" at 200,59 size 25x19; FormatPattern 999
      ProcessValue <- "DB_DTLData_DTL_Imaje Er_1.MINUTE"
   TextField "Text field_3" at 30,42 size 144x17; Text 'Error Counter'
   TextField "Text field_4" at 29,59 size 145x19; Text 'System Imaje Error'
   TextField "Text field_5" at 29,114 size 145x21; Text 'Pressure Low'
   TextField "Text field_6" at 29,133 size 145x20; Text 'Sloft Jammed'
   IOField "I/O field_3" at 175,59 size 25x19; FormatPattern 999
      ProcessValue <- "DB_DTLData_DTL_Imaje Er_1.HOUR"
   TextField "Text field_13" at 196,58 size 8x17; Text ':'
   TextField "Text field_14" at 196,113 size 8x17; Text ':'
   TextField "Text field_15" at 196,133 size 8x17; Text ':'
   TextField "Text field_17" at 220,58 size 8x17; Text ':'
   TextField "Text field_18" at 220,113 size 8x17; Text ':'
   TextField "Text field_19" at 220,133 size 8x17; Text ':'
   TextField "Text field_23" at 196,75 size 8x17; Text ':'
   TextField "Text field_24" at 220,75 size 8x17; Text ':'
   TextField "Text field_26" at 196,93 size 8x17; Text ':'
   TextField "Text field_27" at 220,93 size 8x17; Text ':'

